   // ---------------------------------
   // Simulation

   // IO-mapping for the valves most be commented-out, to make simulation work.
   #motorValveSimulation_1(speed := #speed, io := #valve1.hmi.io);
   #motorValveSimulation_2(speed := #speed, io := #valve2.hmi.io);
END_FUNCTION_BLOCK

FUNCTION_BLOCK "pulsValve"   // FB13, SCL
{ S7_Optimized_Access := 'TRUE' }
VERSION : 0.1
   VAR_INPUT
      iOpening : Bool;
      iCloses : Bool;
      iPuls : Bool;
      iFullyOpen : Bool;
      iFullyClosed : Bool;
      iConfTimeout : Time := T#3S;
      iConfPulsesBetweenOpenAndClosed : Int;
   END_VAR
   VAR_OUTPUT
      qPos : Real;
      qUnknownPos : Bool;
   END_VAR
   VAR
      cnt : Int;
      rtrig_puls : R_TRIG;
      "timer" : IEC_TIMER;
      first_scan : Bool := TRUE;
   END_VAR
   VAR CONSTANT
      NUMBER_PULES_NOT_CONFIGERED : Int := 0;
   END_VAR
BEGIN
   // Valve position based on puls feedback 

   #rtrig_puls(CLK := #iPuls);
   #"timer".TON(IN := (#iOpening OR #iCloses) AND NOT #rtrig_puls.Q,
              PT := #iConfTimeout);
   IF #iConfPulsesBetweenOpenAndClosed = 0 // Number of pules not configured
       OR #"timer".Q
       OR #first_scan  // 
   THEN
       #qUnknownPos := true;
   ELSIF #iFullyOpen THEN
       #cnt := #iConfPulsesBetweenOpenAndClosed;
       #qUnknownPos := false;
   ELSIF #iFullyClosed THEN
       #cnt := 0;
       #qUnknownPos := false;
   ELSE
       IF #iOpening AND #iCloses THEN
           ; // No action
       ELSIF #rtrig_puls.Q THEN
           #cnt += BOOL_TO_INT(#iOpening);
           #cnt -= BOOL_TO_INT(#iCloses);
       END_IF;
   END_IF;
   #qPos := INT_TO_REAL(#cnt) / INT_TO_REAL(#iConfPulsesBetweenOpenAndClosed) * 100;
   #first_scan := false;
END_FUNCTION_BLOCK

FUNCTION_BLOCK "_loadBalancer_example"   // FB14, SCL
{ S7_Optimized_Access := 'TRUE' }
VERSION : 0.1
   VAR
      load_balancer : "loadBalancer";
   END_VAR
   VAR RETAIN
      devices : Array[1..3] of "load_balancer_device_udt";
      settings : "load_balancer_settings_udt";   // Comman settings
   END_VAR
   VAR
      ___ : Bool;
      pid_output : Real;
      in_1_available : Bool;
      in_1_in_opreation : Bool;
      in_2_available : Bool;
      in_2_in_opreation : Bool;
      in_3_available : Bool;
      in_3_in_opreation : Bool;
      out_1 : Bool;
      out_2 : Bool;
      out_3 : Bool;
      out_1_value : Real;
      out_2_value : Real;
      out_3_value : Real;
   END_VAR
BEGIN
   // Load balancer example:

   // - If devices (eg. pumps) work in parallell, the function will add
   //   or remove devices to operate as the demand increase or decrease.
   // - For vfd, there should be configured a long enough ramp time to
   //   make a smooth transition when a device is added or removed for
   //   operation.
   // - More devices can be controlled, by expand the #devices array.
   // - For this theoretically example static variables bellow "___"
   //   are used, in real application the static variables would be
   //   fysical io.

   // - IMPORTANT: both #devices and #settings need to be set to retain.

   // Available: Eg. in auto, no emergensy stop, no comm.error, ready, etc.
   #devices[1].available := #in_1_available;
   #devices[2].available := #in_2_available;
   #devices[3].available := #in_3_available;

   // input:     Typically the output of a pid-controller, the "damand".
   // devices:   A array, one element for each device.
   // settings:  Can be connected to faceplate in hmi, 
   #load_balancer(input := #pid_output,
                  devices := #devices,
                  settings := #settings );
   // - Important: both #devices and #settings need to be set to retain.
   // - Open the block to see the description inside.

   // Output to devices.
   #out_1 := #devices[1].Q;
   #out_2 := #devices[2].Q;
   #out_3 := #devices[3].Q;

   // If vfd devices is controll by a vfd, then the pid_output shuld be forwared
   // to the vfd's:    
   #out_1_value := SEL(G := #devices[1].Q, IN0 := 0, IN1 := #pid_output);
   #out_2_value := SEL(G := #devices[2].Q, IN0 := 0, IN1 := #pid_output);
   #out_3_value := SEL(G := #devices[3].Q, IN0 := 0, IN1 := #pid_output);
END_FUNCTION_BLOCK

FUNCTION_BLOCK "analogIn_fb"   // FB18, SCL
{ S7_Optimized_Access := 'TRUE' }
VERSION : 0.1
   VAR_INPUT
      in : Int;
   END_VAR
   VAR RETAIN
      aiUdt : "analogInUdt";
   END_VAR
   VAR
      normX : "normXAnalogUdt";
   END_VAR
BEGIN

   "analogIn"(in := #in, aiUdt := #aiUdt, normX := #normX);
END_FUNCTION_BLOCK

FUNCTION_BLOCK "example_stateMachine"   // FB21, SCL
{ S7_Optimized_Access := 'TRUE' }
VERSION : 0.1
   VAR
      state : Int;
      timer1 : "stateMachineTimer";
      timer2 : "stateMachineTimer";
      __condition_1__ : Bool := TRUE;
      __condition_2__ : Bool := TRUE;
      HMI_status : String[100];
   END_VAR
BEGIN
   // State machine with timer example. (https://github.com/rexhip/)

   CASE #state OF
       0:  // Next state after 14 sec. Note that the timer is only one line of code.
           #state += BOOL_TO_INT("sTimer"(pt := T#14s, t := #timer1));

           #HMI_status := CONCAT(IN1 := 'State 0, remaining time: ',
                                 IN2 := "::"(in := #timer1.rt), IN3 := '.');

       1:  // Next state after 7 sec, and '__condition_1__' is true.
           #timer1.pt := T#7s;
           #state += BOOL_TO_INT(#timer1.q AND #__condition_1__);

           // Back to stae 0 if 50 sec elapses. A timer can be used once in each state,
           // therfor timer2 used for this condition. Note the ":=" and not "+=" as above.
           #state := SEL(G := "sTimer"(pt := T#1m50s, t := #timer2), IN0 := #state, IN1 := 0);

           #HMI_status := CONCAT(IN1 := 'State 1, Timer1 ', IN2 := "::"(in := #timer1.rt),
                                 IN3 := ', Timer2 ', IN4 := "::"(in := #timer2.rt));

       2:  // Back to state 0, when '__condition_2__' has been true for 8 sec continuously.
           // The sTimer FC could have been used here also, but for the sake of the
           // example it isn't.
           IF #__condition_2__ THEN
               #timer1.pt := T#8s;
               #state := SEL(G := #timer1.q, IN0 := #state, IN1 := 0);
           END_IF;

           #HMI_status := 'State 2.';
   END_CASE;

   #timer1(state := #state); // Run the timer code.
   #timer2(state := #state);
END_FUNCTION_BLOCK

FUNCTION_BLOCK "modbus_test_rtu_1500"   // FB102, SCL
{ S7_Optimized_Access := 'TRUE' }
VERSION : 0.1
   VAR
      mb_master_1500_ctrl : "mb_master_1500_ctrl";
      mb_query : "mb_query";
      temperature_1 : "Jdrk_RS_WS_N01_8";
      temperature_2 : "Jdrk_RS_WS_N01_8";
      temperature_3 : "Jdrk_RS_WS_N01_8";
      sb_temp_no_answer_1 : "sb_temp_no_answer";
      sb_temp_no_answer_2 : "sb_temp_no_answer";
      sb_temp_no_answer_3 : "sb_temp_no_answer";
      sb_temp_error_1 : "sb_temp_error";
      sb_temp_error_2 : "sb_temp_error";
      sb_temp_error_3 : "sb_temp_error";
      delay_between_queries : "mb_delay_between_queries";
      mb_delay : "mb_delay";
   END_VAR
BEGIN

   #mb_master_1500_ctrl.conf.parity := 0;
   #mb_master_1500_ctrl(hardware_id := 269,
                        operating_mode := 4,
                        baud := 9600,
                        mb_query := #mb_query);

   #delay_between_queries(mb_query := #mb_query);


   #temperature_1(mb_query := #mb_query);
   #temperature_2(mb_query := #mb_query);
   #temperature_3(mb_query := #mb_query);

   #mb_delay(mb_query := #mb_query);

   #sb_temp_no_answer_1(mb_query := #mb_query);
   #sb_temp_no_answer_2(mb_query := #mb_query);
   #sb_temp_no_answer_3(mb_query := #mb_query);

   #sb_temp_error_1(mb_query := #mb_query);
   #sb_temp_error_2(mb_query := #mb_query);
   #sb_temp_error_3(mb_query := #mb_query);
END_FUNCTION_BLOCK

FUNCTION "movingAverageFilter" : Void   // FC1, SCL
{ S7_Optimized_Access := 'TRUE' }
VERSION : 0.1
   VAR_INPUT
      in : Real;
   END_VAR
   VAR_IN_OUT
      filterConst : Real;   // 0=off.
      Q : Real;
   END_VAR
   VAR_TEMP
      z : LReal;
   END_VAR
BEGIN
   // Running average smoothing filter.
   //  - Filter constant has to greater then zero
   //  - PLC scan time will affect the filter.

   IF #filterConst = 0 THEN // Zero -> disable filter 
       #Q := #in;
   ELSE
       #filterConst := MAX(IN1 := 0, IN2 := #filterConst);
       // Creating a number betwwen zero and less then one.
       #z := -1 / REAL_TO_LREAL(#filterConst + 1); 
       #Q := LREAL_TO_REAL(#z * REAL_TO_LREAL(#Q)
                           + (1 - #z) * REAL_TO_LREAL(#in));
   END_IF;
END_FUNCTION

FUNCTION "real2time_format" : Time   // FC1, SCL
{ S7_Optimized_Access := 'TRUE' }
VERSION : 0.1
   VAR_INPUT
      in : Real;
      format : SInt;   // 1=ms, 2=sec, 3=min, 4=h, 5=day
   END_VAR
BEGIN
   // PT-max: 24 days, 20 hours, 31 min, 23 sec and 647 ms.

   // Format: 1=ms, 2=sec, 3=min, 4=h, 5=day

   #real2time_format := T#0s;
   CASE #format OF
       1:  // ms
           #real2time_format := T_CONV(REAL_TO_DINT(#in));
       2:  // Sec
           #real2time_format := T_CONV(REAL_TO_DINT(#in * 1000));
       3:  // Min
           #real2time_format := T_CONV(REAL_TO_DINT(#in * 60000)); //  1000*60
       4:  // Hours
           #real2time_format := T_CONV(REAL_TO_DINT(#in * 3600000)); // 1000*60*60
       5:  // Days
           #real2time_format := T_CONV(REAL_TO_DINT(#in * 86400000)); // 1000*60*60*24
   END_CASE;
END_FUNCTION

FUNCTION "time2real_format" : Real   // FC2, SCL
{ S7_Optimized_Access := 'TRUE' }
VERSION : 0.1
   VAR_INPUT
      in : Time;
      format : SInt;   // 1=ms, 2=sec, 3=min, 4=h, 5=day
   END_VAR
BEGIN
   // PT-max: 24 days, 20 hours, 31 min, 23 sec and 647 ms.

   // Format: 1=ms, 2=sec, 3=min, 4=h, 5=day

   #time2real_format := 0;
   CASE #format OF
       1:  // ms
           #time2real_format := DINT_TO_REAL(T_CONV(#in));
       2:  // Sec
           #time2real_format := DINT_TO_REAL(T_CONV(#in)) / 1000;
       3:  // Min
           #time2real_format := DINT_TO_REAL(T_CONV(#in)) / 60000; // 1000*60
       4:  // Hours
           #time2real_format := DINT_TO_REAL(T_CONV(#in)) / 3600000; // 1000*60*60
       5:  // Days
           #time2real_format := DINT_TO_REAL(T_CONV(#in)) / 86400000; // 1000*60*60*24
   END_CASE;
END_FUNCTION

FUNCTION "analogIn" : Void   // FC4, SCL
TITLE = Analog input
{ S7_Optimized_Access := 'TRUE' }
VERSION : 0.1
   VAR_INPUT
      in : Int;
   END_VAR
   VAR_IN_OUT
      aiUdt : "analogInUdt";
      normX : "normXAnalogUdt";
   END_VAR
   VAR_TEMP
      u : Real;
      x : Real;
      y : Real;
      "e" : Int;
   END_VAR
BEGIN
   // Analog input scaling.

   #u := NORM_X(MIN := #normX.rawMin, VALUE := #in, MAX := #normX.rawMax);
   "movingAverageFilter"(in := #u,
                         filterConst := #aiUdt.filterConst,
                         Q := #aiUdt.unitInterval);
   IF #aiUdt.sim THEN
       ; // A simulated value can be set directly to #aiUdt.Q and #aiUdt.Error
   ELSE
       // Scale back up to raw-value to check if outside error limits.
       #x := SCALE_X(MIN := #normX.rawMin, MAX := #normX.rawMax,
                     VALUE := #aiUdt.unitInterval);
       #aiUdt.Error := #x < #normX.errorLimMin OR #x > #normX.errorLimMax;
       // Log the time when the error occurred.
       IF #aiUdt.Error AND NOT #aiUdt.zOldError THEN
           #"e" := RD_LOC_T(#aiUdt.ErrorTime);
       END_IF;

       IF #aiUdt.Error THEN
           #y := SINT_TO_REAL(#aiUdt.errorAction) / 100;
       ELSIF #aiUdt.forceInsideScale THEN
           #y := LIMIT(MN := 0, IN := #aiUdt.unitInterval, MX := 1);
       ELSE
           #y := #aiUdt.unitInterval;
       END_IF;
       #aiUdt.Q := SCALE_X(MIN := #aiUdt.scaleMin, MAX := #aiUdt.scaleMax,
                           VALUE := #y ) * #aiUdt.gain + #aiUdt.offset;
   END_IF;
   #aiUdt.zOldError := #aiUdt.Error;

   // ( https://github.com/rexhip/ )
END_FUNCTION

FUNCTION "boost_start" : Void   // FC5, SCL
{ S7_Optimized_Access := 'TRUE' }
VERSION : 0.1
   VAR_INPUT
      t_diff : USInt;
      start : Bool;
   END_VAR
   VAR_OUTPUT
      reset_timers : Bool;
   END_VAR
   VAR_IN_OUT
      devices : Array[*] of "load_balancer_device_udt";
      settings : "load_balancer_settings_udt";
      info : "load_balancer_info_udt";
      boost_start : SInt;
      set : SInt;
   END_VAR
   VAR_TEMP
      c : DInt;
      u : DInt;
      lower : DInt;
   END_VAR
BEGIN
   #lower := LOWER_BOUND(ARR := #devices, DIM := 1);
   FOR #c := #lower TO UPPER_BOUND(ARR := #devices, DIM := 1) DO

       #u := #c - #lower + 1; // #u start at 1, increasing by 1 for each iteration.
       IF #settings.boostStart.reset THEN
           // Reset stastic, on how many devices is operating same time.
           #devices[#c].z.n_cnt := 0;
       ELSIF #settings.info.started = #u THEN
           // Log how many devices is operating same time, most fequently.
           #devices[#c].z.n_cnt += #t_diff;
       END_IF;

       // Change how many devices to boost start at startup, based on how many
       // devices is most commenly used.
       IF #settings.boostStart.auto
           AND #devices[#c].z.n_cnt >
           (* *)#devices[#lower + #settings.boostStart.devices - 1].z.n_cnt
       THEN
           #settings.boostStart.devices := DINT_TO_USINT(#u);
       END_IF;
   END_FOR;

   // Set a number of operating devices. (Without waiting for the input and the timers)
   IF #set > -1 THEN
       #boost_start := #set - UINT_TO_SINT(#info.devices_started);

       // Do boost start when input change away from zero.    
   ELSIF #settings.boostStart.enable // HMI enable.
       AND #start
       AND #set = -1
   THEN
       #boost_start :=
       UINT_TO_SINT(#settings.boostStart.devices - #info.devices_started);
   END_IF;
   // #set is put back to -1 at the bottom of the block.

   // MN: Devies started to be stopped.
   // MX: Devices available for start. 
   #boost_start := LIMIT(MN := - UINT_TO_SINT(#info.devices_started),
                         IN := #boost_start,
                         MX := UINT_TO_SINT(#info.devices_standby));

   #reset_timers := #boost_start <> 0 OR #set <> -1; // Reset timers.
END_FUNCTION

FUNCTION "analogInReal" : Void   // FC7, SCL
{ S7_Optimized_Access := 'TRUE' }
VERSION : 0.1
   VAR_INPUT
      in : Real;
      error : Bool;
   END_VAR
   VAR_IN_OUT
      aiUdt : "analogInAndAlarmsUdt";
      ioGlobal : "ioGlobal_FB";
   END_VAR
   VAR_TEMP
      dommy : Int;
      u : Real;
   END_VAR
BEGIN
   // Analog input 
   // Wrapper to use analog input block with real input.
   // 
   #aiUdt.ai.Error := #error;

   IF #aiUdt.ai.sim THEN
       ; // A simultated value may be set directly at: #ai.ai.Q
   ELSE
       #u := #in * #aiUdt.ai.gain + #aiUdt.ai.offset;
       "movingAverageFilter"(in := #u,
                             filterConst := #aiUdt.ai.filterConst,
                             Q := #aiUdt.ai.Q);
   END_IF;

   #aiUdt.execAiLogic := false;
   "analogInAndAlarms"(in := #dommy,
                       aiUdt := #aiUdt,
                       ioGlobal := #ioGlobal);

   // ( https://github.com/rexhip/ )
END_FUNCTION

FUNCTION "analogOut" : Void   // FC9, SCL
{ S7_Optimized_Access := 'TRUE' }
VERSION : 0.1
   VAR_OUTPUT
      q : Int;
   END_VAR
   VAR_IN_OUT
      aoUdt : "analogOutUdt";
      ioGlobal : "ioGlobal_FB";
   END_VAR
   VAR_TEMP
      x : Real;
      y : Real;
   END_VAR
BEGIN
   // Analog out 

   // - failSafe: Output will go to a predefined value set by
   //   failSafeValue (%), this can be used for emergency stop.
   //   Simulation will not work when failSafe is activated.

   // A id for each io
   #ioGlobal.z.ioIdCnt += 1;

   IF #ioGlobal.info2ioBlocks.disableAllSim THEN
       #aoUdt.simEnable := false;
   END_IF;

   IF #aoUdt.failSafe THEN
       #x := SINT_TO_REAL(#aoUdt.failSafeValue) / 100 ; // [%]
   ELSE
       IF #aoUdt.simEnable THEN
           #y := #aoUdt.simValue;
       ELSIF #aoUdt.interlook THEN
           #y := 0;
       ELSE
           #y := #aoUdt.in;
       END_IF;
       #x := NORM_X(MIN := #aoUdt.scaleMin, VALUE := #y,
                    MAX := #aoUdt.scaleMax);
       #aoUdt.simValue := #y;
   END_IF;
   #x := LIMIT(MN := 0, IN := #x, MX := 1);
   #q := SCALE_X(MIN := #ioGlobal.normX.rawMin, VALUE := #x,
                     MAX := #ioGlobal.normX.rawMax);

   #ioGlobal.collectInfo.activeSimCnt += BOOL_TO_UINT(#aoUdt.simEnable);

   // ( https://github.com/rexhip/ )
END_FUNCTION

FUNCTION "ioGlobalMotorValveLinking" : Void   // FC24, SCL
{ S7_Optimized_Access := 'TRUE' }
VERSION : 0.1
   VAR_IN_OUT
      ioGlobal : "ioGlobal_FB";
      valve : "motorValve";
   END_VAR
BEGIN
   // Link ioGlobal with valve functions.

   // A id for each io
   #ioGlobal.z.ioIdCnt += 1;

   IF #ioGlobal.info2ioBlocks.disableAllSim THEN
       #valve.hmi.sim.enable := false;
   END_IF;
   // Count active simulations
   #ioGlobal.collectInfo.activeSimCnt +=
   BOOL_TO_UINT(#valve.hmi.sim.enable OR #valve.hmi.sim.simByPlc);

   // Count number of errors
   #ioGlobal.collectInfo.errorCnt +=
   BOOL_TO_UINT(#valve.hmi.io.in.posError OR #valve.hmi.error.timeout);
END_FUNCTION

FUNCTION "real_to_time" : Time   // FC29, SCL
{ S7_Optimized_Access := 'TRUE' }
VERSION : 0.1
   VAR_INPUT
      in : Real;
   END_VAR
BEGIN

   #real_to_time := T_CONV(REAL_TO_DINT(#in * 1000));
END_FUNCTION

// folder: Library/Alternating/Load balancer/Blocks and UDT's

FUNCTION_BLOCK "loadBalancer"   // FB13, SCL
{ S7_Optimized_Access := 'TRUE' }
VERSION : 0.1
   VAR_INPUT
      input : Real;   // [%] Typically a output from a pid-controller.
   END_VAR
   VAR_IN_OUT
      devices : Array[*] of "load_balancer_device_udt";   // Variables for each device.
      settings : "load_balancer_settings_udt";   // Comman settings
   END_VAR
   VAR RETAIN
      conf : Struct   // Advanced configuration
         enable_operation_time_cnt : Bool := true;   // Enable operation time cnt
         at_least_one : Bool := true;   // At least one device will always be in operation
         bypass_InOperation_signal : Bool := true;   // Output control in-operation variable.
         input_zero_reset : Time := T#10M;   // All outputs will be turn off if input has been zero for this time.
         exec_boost_start_code : Bool := true;
      END_STRUCT;
   END_VAR
   VAR
      boost_start : SInt;   // Start a relative number of devices. (Negative number will stop devices)
      set : SInt := -1;   // Start a exact number of devices. (Set back to -1 right away)
      _ : Bool;
      timer_start : IEC_TIMER;
      timer_start_q : Bool;
      timer_stop : IEC_TIMER;
      timer_stop_q : Bool;
      timer_input_zero : IEC_TIMER;
      old_sec : USInt;
      ftrig_zero_input_timer : F_TRIG;
      runtime_mem1 : LReal;
      runtime_mem2 : LReal;
   END_VAR
   VAR_TEMP
      candidates : Struct
         start : Struct
            index : DInt;
            operation_time : UDInt;
         END_STRUCT;
         stop : Struct
            index : DInt;
            operation_time : UDInt;
         END_STRUCT;
      END_STRUCT;
      info : "load_balancer_info_udt";
      lower : DInt;
      upper : DInt;
      c : DInt;
      t_diff : USInt;
      oper : SInt;
      u : DInt;
      reset_timers : Bool;
      dommy : Bool;
   END_VAR
   VAR CONSTANT
      NO_CANDIDATE : DInt := 16#7fffffff;
   END_VAR
BEGIN
   (* === Load balancer ===    

   - If devices (eg. pumps) work in parallell, the function will start or stop devices
     to operate as the demand increase or decrease.
   - A devices will be added for operation, if #input is above a certain value for a
     ceratin time, eg above 90% for 50 seconds. Likewise a devices will be removed from
     operation if #input is bellow a certain value for a certain time, eg. 10% for 30
     secunds. The limits and the times are adjustable inside #settings.
   - It's the device with least operating time that will be added first, and the device
     with most operating hours will be removed from operation first.
   - #input will typically be the output of a pid-controller.
   - For vfd, there should be configured a ramp time to make a smooth transition when a
     device is added or removed for operation.
   - #devices[*].in.in_operation, is a input for fyscical feedback signal from the
     devices. this feature can be disabled by setting
     #load_balancer.conf.bypass_InOperation_signal, to true.
   - #boost_start: Make more then one devices start right away, without have to wait for
     them to start one by one. Use a negative number to stop several devies at once. One
     scan is need to start or stop each device.
   - #set: Will start or stop devies to mache number of the variable. This block will set
     the variable to -1 for the next scan.

   *)

   // If input is zero for a certain time, then all outputs is set to false.
   #timer_input_zero.TON(IN := #input = 0, PT := #conf.input_zero_reset);
   // Used to set correct number of devices from start. (Boost start)
   #ftrig_zero_input_timer(CLK := NOT #timer_input_zero.Q);

   // Default values, if the value isn't overwritten after the
   // for-loop (bellow), then there is "no candidate".
   #candidates.stop.index := #NO_CANDIDATE;
   #candidates.start.index := #NO_CANDIDATE;
   // Set to max, try find a lesser value in the for-loop bellow.
   #candidates.start.operation_time := 16#ffffffff;

   // Operating time preparing calculations:
   #runtime_mem2 += RUNTIME(#runtime_mem1);
   #t_diff := LREAL_TO_USINT(FLOOR(#runtime_mem2)); // "Overflow" if >= 1 sec.
   #runtime_mem2 -= USINT_TO_LREAL(#t_diff);

   // Boost start makes, more then one device start right away.
   IF #conf.exec_boost_start_code THEN
       "boost_start"(t_diff := #t_diff,
                     start := #ftrig_zero_input_timer.Q,
                     reset_timers => #reset_timers,
                     devices := #devices,
                     settings := #settings,
                     info := #info,
                     boost_start := #boost_start,
                     set := #set);
   END_IF;

   #lower := LOWER_BOUND(ARR := #devices, DIM := 1);
   #upper := UPPER_BOUND(ARR := #devices, DIM := 1);
   FOR #c := #lower TO #upper DO

       #devices[#c].Q := #devices[#c].Q
       (* *)AND #devices[#c].available // Disable devices that are not available. 
       (* *)AND NOT #timer_input_zero.Q // Input has not been zero for a ceratain time.
       OR #settings.bypass; // If bypass, then enable all devices.

       // If no fysical feedback signal from device for "in-operation", then
       // it's possible to bypass it.
       IF #conf.bypass_InOperation_signal THEN
           #devices[#c].in_operation := #devices[#c].Q;
       END_IF;

       REGION Candidates        
           // Candidate device to be stoped (the one that has the longest operating time)
           IF #devices[#c].Q // In use
               AND #devices[#c].operation_time >= #candidates.stop.operation_time
           THEN
               #candidates.stop.index := #c;
               #candidates.stop.operation_time := #devices[#c].operation_time;
           END_IF;

           // Candidate device to be started (the one that has the least operating time)
           IF #devices[#c].available
               AND NOT #devices[#c].Q // not allready in use
               AND #devices[#c].operation_time < #candidates.start.operation_time
           THEN
               #candidates.start.index := #c;
               #candidates.start.operation_time := #devices[#c].operation_time;
           END_IF;
       END_REGION

       REGION Collect-statistics
           // Operating time cnt. (#t_diff will always be zero, if the feature is disabled)
           #devices[#c].operation_time += SEL(G := #devices[#c].in_operation
                                              AND #conf.enable_operation_time_cnt,
                                              IN0 := 0, IN1 := USINT_TO_UDINT(#t_diff));
           // Count number of devices in operation.
           #info.devices_in_operation += BOOL_TO_UINT(#devices[#c].in_operation);
           // Count number of devices in standby.
           #info.devices_standby +=
           BOOL_TO_UINT(#devices[#c].available
                        AND NOT #devices[#c].Q); // NOT #devices[#c].in.in_operation
           // Count number of devices started.
           #info.devices_started += BOOL_TO_UINT(#devices[#c].Q);
       END_REGION
   END_FOR;

   // Some info (for hmi)
   #settings.info.total := DINT_TO_UINT(#upper - #lower + 1);

   // If for some reason, the number operating devies can be limited to less
   // then available
   #settings.max_devices_same_time := // A setting.
   LIMIT(MN := 1,
         IN := #settings.max_devices_same_time,
         MX := #settings.info.total);

   // Force min value for param.
   #settings.max_diff_operating.sec :=
   MAX(IN1 := 60, IN2 := #settings.max_diff_operating.sec);

   // Timers for adding and removing devices for operation.

   #timer_stop.TON(IN := #input < #settings.stop.limit AND NOT #reset_timers,
                   PT := #settings.stop.delay,
                   Q => #timer_stop_q);
   #timer_start.TON(IN := #input > #settings.start.limit AND NOT #reset_timers,
                    PT := #settings.start.delay,
                    Q => #timer_start_q);

   REGION start-stopp
       // Stoping a device
       IF NOT #settings.bypass // The bypass-function turn on all outputs. 
           AND #candidates.stop.index <> #NO_CANDIDATE // A device is available 
           AND (#info.devices_in_operation > 1 // Can't remove last device in operation
           (* *)OR NOT #conf.at_least_one)  // Possible to disable the feature
           AND (
           (* *)#info.devices_in_operation > #settings.max_devices_same_time
           (* *)OR #timer_stop_q // If #input below a certain value for a certain time
           (* *)OR #settings.stop.force  // Used to stop the next device (hmi)
           (* *)OR #boost_start < 0)
       THEN
           #devices[#candidates.stop.index].Q := false; // Disable one device
           RESET_TIMER(#timer_stop);
           #oper := -1;
           // Increase var until zero.
           #boost_start := SEL(G := #boost_start < 0, IN0 := 0, IN1 := #boost_start + 1);

           // Start a devices.
       ELSIF #candidates.start.index <> #NO_CANDIDATE // A device is available 
           AND #info.devices_in_operation < #settings.max_devices_same_time
           AND #input > 0 AND (
           (* *)#info.devices_in_operation < 1 // At least one device operating
           (*      *)AND #conf.at_least_one // Possible to disable the feature
           (* *)OR #timer_start_q // If #input above a certain value for a certain time
           (* *)OR #settings.start.force // Used to starp the next device (hmi)
           (* *)OR #boost_start > 0)
       THEN
           #devices[#candidates.start.index].Q := true; // Enable one more device
           RESET_TIMER(#timer_start);
           #oper := 1;
           // Decrease var until zero.
           #boost_start := SEL(G := #boost_start > 0, IN0 := 0, IN1 := #boost_start - 1);

           // Change operating device, if the operating-time between two devies is to large.
       ELSIF #settings.max_diff_operating.enable
           AND #candidates.start.index <> #NO_CANDIDATE // A candidate is available to be started
           AND #candidates.stop.index <> #NO_CANDIDATE // A candidate is available to be stoped
           AND (#candidates.stop.operation_time - #candidates.start.operation_time >
           (* *)#settings.max_diff_operating.sec) // And the difference is to large.
       THEN
           // Stop the device with most operating time and start the devices with
           // least operating time.
           #devices[#candidates.stop.index].Q := false;
           #devices[#candidates.start.index].Q := true;
       END_IF;
   END_REGION

   // Update vars, after start or stop a device. (above)
   #info.devices_in_operation += SINT_TO_UINT(#oper);
   #info.devices_started += SINT_TO_UINT(#oper);
   #info.devices_standby -= SINT_TO_UINT(#oper);

   // Transfer values to hmi-vars
   #settings.info.in_operation := #info.devices_in_operation;
   #settings.info.started := #info.devices_started;
   #settings.info.standby := #info.devices_standby;

   #settings.info.input := #input;

   // Information has been recived, so now back to default values.
   #set := -1;
   #settings.start.force := false;
   #settings.stop.force := false;
   #settings.boostStart.reset := false;

   // https://github.com/rexhip/
END_FUNCTION_BLOCK

// folder: Library/IO-handeling/Analog in/Blocks

FUNCTION "analogInAndAlarms" : Void   // FC6, SCL
{ S7_Optimized_Access := 'TRUE' }
VERSION : 0.1
   VAR_INPUT
      in : Int;
   END_VAR
   VAR_IN_OUT
      aiUdt : "analogInAndAlarmsUdt";
      ioGlobal : "ioGlobal_FB";
   END_VAR
   VAR CONSTANT
      VALUE_LESS_THEN_LIM : SInt := 1;
      VALUE_GREATER_THEN_LIM : SInt := 2;
   END_VAR
BEGIN
   // Analog input with alarm handling. 

   REGION Input handling
       // A id for each io
       #ioGlobal.z.ioIdCnt += 1;

       // Disable all simulations.
       #aiUdt.ai.sim := #aiUdt.ai.sim AND NOT #ioGlobal.info2ioBlocks.disableAllSim;

       IF #aiUdt.execAiLogic THEN // Execute analog input logic
           "analogIn"(in := #in,
                      aiUdt := #aiUdt.ai,
                      normX := #ioGlobal.normX);
       END_IF;
       // Count number of errors
       #ioGlobal.collectInfo.errorCnt += BOOL_TO_UINT(#aiUdt.ai.Error);;
       // Count active simulations 
       #ioGlobal.collectInfo.activeSimCnt += BOOL_TO_UINT(#aiUdt.ai.sim);
   END_REGION

   REGION Alarms  
   // Connecting ioGlobal functions with each alarm.
   "ioGlobalAlarmLinking"(alarm := #aiUdt.alarmHH, ioGlobal := #ioGlobal);
   "ioGlobalAlarmLinking"(alarm := #aiUdt.alarmH, ioGlobal := #ioGlobal);
   "ioGlobalAlarmLinking"(alarm := #aiUdt.alarmLL, ioGlobal := #ioGlobal);
   "ioGlobalAlarmLinking"(alarm := #aiUdt.alarmL, ioGlobal := #ioGlobal);

   "alarmReal"(value := #aiUdt.ai.Q, // HH alarm
               action := #VALUE_GREATER_THEN_LIM,
               disable := false,
               runtimeDiff := #ioGlobal.info2ioBlocks.runtimeDiff,
               alarm := #aiUdt.alarmHH);
   "alarmReal"(value := #aiUdt.ai.Q,// H alarm
               action := #VALUE_GREATER_THEN_LIM,
               disable := #aiUdt.alarmHH.Q,
               runtimeDiff := #ioGlobal.info2ioBlocks.runtimeDiff,
               alarm := #aiUdt.alarmH);
   "alarmReal"(value := #aiUdt.ai.Q, // LL alarm
               action := #VALUE_LESS_THEN_LIM,
               disable := false,
               runtimeDiff := #ioGlobal.info2ioBlocks.runtimeDiff,
               alarm := #aiUdt.alarmLL);
   "alarmReal"(value := #aiUdt.ai.Q, // L alarm
               action := #VALUE_LESS_THEN_LIM,
               disable := #aiUdt.alarmLL.Q,
               runtimeDiff := #ioGlobal.info2ioBlocks.runtimeDiff,
               alarm := #aiUdt.alarmL);
   END_REGION

   REGION HMI-features
       // Copy paste all settings. (HMI)
       IF #aiUdt.hmi.copyAllSettings THEN
           #ioGlobal.copyPaste := #aiUdt;
           #aiUdt.hmi.copyAllSettings := false;
       ELSIF #aiUdt.hmi.pasteAllSettings THEN
           "pasteAnalogInSetting"(src := #ioGlobal.copyPaste, dest := #aiUdt);
           #aiUdt.hmi.pasteAllSettings := false;
       END_IF;

       #aiUdt.hmi.showTag := #ioGlobal.hmi.hmiShowTags;
   END_REGION

   // ( https://github.com/rexhip/ )
END_FUNCTION

FUNCTION "analogInSimple" : Real   // FC13, SCL
{ S7_Optimized_Access := 'TRUE' }
VERSION : 0.1
   VAR_INPUT
      mn : Real;
      in : Int;
      mx : Real;
   END_VAR
   VAR_TEMP
      x : Real;
   END_VAR
BEGIN
   // Analog in 

   #x := NORM_X(MIN := 0, VALUE := #in, MAX := 27648);
   #x := LIMIT(MN := 0, IN := #x, MX := 1);
   #analogInSimple := SCALE_X(MIN := #mn, VALUE := #x, MAX := #mx);

   // ( https://github.com/rexhip/ )
END_FUNCTION

// folder: Library/Modbus/.Start examples

FUNCTION_BLOCK "modbus_rtu_1500"   // FB5, SCL
{ S7_Optimized_Access := 'TRUE' }
VERSION : 0.1
   VAR
      mb_query : "mb_query";
      mb_master_1500_ctrl : "mb_master_1500_ctrl";
      abb_aquaMaster_device1 : "abb_aquaMaster_3";
      abb_aquaMaster_device2 : "abb_aquaMaster_3";
      abb_aquaMaster_device3 : "abb_aquaMaster_3";
      resault_data_1 : Word;
   END_VAR
BEGIN
   // hardware_id:     May be found inside the hardware configuration.
   // operating_mode:  0: RS232, 2: RS422, 4: RS485.
   // baud:            Bits per sec. (Parity is even by default)
   // timeout:         Automatically calculated if set to zero. (T#0s)
   // mb_query:        The FB that connects everything together.
   #mb_master_1500_ctrl(hardware_id := 0, // REPLACE WITH CORRECT ID.
                        operating_mode := 4, // RS-485
                        baud := 19200, // bps
                        mb_query := #mb_query);

   // Each blocks bellow represent one device on the bus. 
   #abb_aquaMaster_device1(mb_addr := 1, mb_query := #mb_query);
   #abb_aquaMaster_device2(mb_addr := 2, mb_query := #mb_query);
   #abb_aquaMaster_device3(mb_addr := 3, mb_query := #mb_query);


   // Debugging tip, (no code)
   "mb_Debugging"();
END_FUNCTION_BLOCK

FUNCTION_BLOCK "modbus_tcp"   // FB79, SCL
{ S7_Optimized_Access := 'TRUE' }
VERSION : 0.1
   VAR
      mb_query : "mb_query";
      mb_client_ctrl : "mb_client_ctrl";
      siemens_PAC3200 : "siemens_PAC3200";
      ip : Array[1..4] of Byte;
      mb_delay_between_queries : "mb_delay_between_queries";
   END_VAR
BEGIN
   // IP-address of the modbus server
   #ip[1] := 192;
   #ip[2] := 168;
   #ip[3] := 1;
   #ip[4] := 2;

   // interface:  Profinet interface.
   //             (Find const. inside "Device configuration")
   // conn_id:    A unique id for each tcp connectin in the plc.
   // ip_addr:    The ip-address of the server. (Array of 4 bytes)
   // tcp_port:   Default port is 502. (UDP isn't available)
   // timeout:    Depends on the network conncetion.
   // mb_query:   The query FB.
   #mb_client_ctrl(interface := 0, // REPLACE WITH CORRECT ID OR CONST,
                                   // Eg. "Local~PROFINET_interface_1",
                   conn_id := 123,
                   ip_addr := #ip,
                   tcp_port := 502,
                   timeout := T#400ms,
                   mb_query := #mb_query);

   // Delay the query execution, this prevent the plc from
   // jamming the network. Adjust the time to the application.
   #mb_delay_between_queries(delay := T#500ms,
                             mb_query := #mb_query);

   #siemens_PAC3200(mb_query := #mb_query);


   // Debugging tip, (no code)
   "mb_Debugging"();
END_FUNCTION_BLOCK

FUNCTION_BLOCK "modbus_rtu_1200"   // FB98, SCL
{ S7_Optimized_Access := 'TRUE' }
VERSION : 0.1
   VAR
      mb_query : "mb_query";
      mb_master_1200_ctrl : "mb_master_1200_ctrl";
      abb_aquaMaster_device1 : "abb_aquaMaster_3";
      abb_aquaMaster_device2 : "abb_aquaMaster_3";
      abb_aquaMaster_device3 : "abb_aquaMaster_3";
      Auma_valve : "Auma_valve";
      Phoenix_Contact_UPS : "Phoenix_Contact_UPS";
      resault_data_1 : Word;
      Phoenix_Contact_UPS_1 : "Phoenix_Contact_UPS";
   END_VAR
BEGIN
   // hardware_id: Can be found inside "Device configuration".
   // baud:        Bits per sec. (Parity is even by default)
   // timeout:     Automatically calculated if set to T#0s.
   // mb_query:    The FB that connects everything together.
   #mb_master_1200_ctrl(hardware_id := 0, // REPLACE WITH CORRECT ID.
                        baud := 19200,
                        mb_query := #mb_query);

   // Each blocks bellow represent one device on the bus.

   // Three Abb aqua-master's.
   #abb_aquaMaster_device1(mb_addr := 1, mb_query := #mb_query);
   #abb_aquaMaster_device2(mb_addr := 2, mb_query := #mb_query);
   #abb_aquaMaster_device3(mb_addr := 3, mb_query := #mb_query);

   // A valve 
   #Auma_valve(mb_addr := 4, mb_query := #mb_query);

   // A UPS.
   #Phoenix_Contact_UPS(mb_addr := 5, mb_query := #mb_query);

   // A station block can be used both for both modbus rtu and tcp. This
   // is particular useful if a tcp-rtu-gateway is used. The same program
   // could be used, just swap mb_master_1200_ctrl, with mb_client_ctrl.

   // Read holding register 456 from device with modbus address 123.
   // This is an example showing that a query does not necessarily need
   // to be part of a station block (SB) as obove, however making
   // reusable SB's is good practice.
   #mb_query(mb_addr := 123,
             mode := #mb_query.c.read.holding_reg,
             data_addr := 456,
             data_ptr := #resault_data_1);


   // Debugging tip, (no code)
   "mb_Debugging"();
END_FUNCTION_BLOCK

FUNCTION "mb_Readme" : Void   // FC13, SCL
{ S7_Optimized_Access := 'TRUE' }
VERSION : 0.1
BEGIN
   (* Instructions:

   - Add one of the exmple FB's to your PLC.
   - Call that FB from a cyclic OB.
   - Terminate connection to type on the example FB. (Right click the FB)
   - Set hardware_id, buad-rate, ip, tcp-port, etc, to the correct value.
   - Look inside the library and check if there is a ready station block (SB),
     for your program. If there isn't then a new has to be made. 
   - Station blocks can be single-DB's or multi-instances in a FB.
   - Remove the exmple code and example SB's.

   IMPORTANT: As stated above, the start examples fb, need to be terminated 
              from it's type. If the type is edited and later there is a 
              library update, then all the changes will get lost.

   - Instructions need to be of the latest version, 
     this is usually already set:
     * Instructions -> Communication -> Others -> Modbus TCP
     * Instructions -> Communication -> Communication processor -> Modbus
     * Instructions -> Communication -> Communication processor -> Modbus (RTU)  
     * Instructions -> Basic instructions -> Word logic operations -> SEL.
     Change version in the right column.

   *)
END_FUNCTION

// folder: Library/Modbus/.Start examples/Other start examples

FUNCTION_BLOCK "LAD_modbus_rtu"   // FB97, LAD
TITLE = Example modbus rtu
{ S7_Optimized_Access := 'TRUE' }
VERSION : 0.1
// REPLACE hardware_id WITH CORRECT ID.
   VAR
      mb_master_ctrl : "mb_master_1200_ctrl";
      mb_query : "mb_query";
      aquaMaster_device1 : "abb_aquaMaster_3";
      aquaMaster_device2 : "abb_aquaMaster_3";
      Auma_valve : "Auma_valve";
      Phoenix_Contact_UPS : "Phoenix_Contact_UPS";
   END_VAR
   VAR_TEMP   // added for the SCL form of the ladder/FBD networks
      _w1 : Bool;
   END_VAR
BEGIN

REGION Network 1: Modbus master
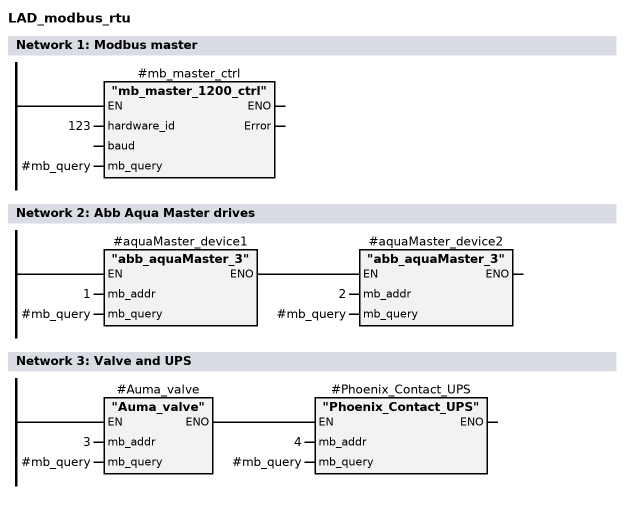
   RUNG wire#powerrail
      #mb_master_ctrl(hardware_id := 123, baud :=, mb_query := #mb_query, Error =>)
   END_RUNG
   // the same network as SCL:
   #mb_master_ctrl(hardware_id := 123, mb_query := #mb_query);   // "mb_master_1200_ctrl"
END_REGION

REGION Network 2: Abb Aqua Master drives
   RUNG wire#powerrail
      #aquaMaster_device1(mb_addr := 1, mb_query := #mb_query)
      #aquaMaster_device2(mb_addr := 2, mb_query := #mb_query)
   END_RUNG
   // the same network as SCL:
   #aquaMaster_device1(mb_addr := 1, mb_query := #mb_query, ENO => #_w1);   // "abb_aquaMaster_3"
   IF #_w1 THEN
       #aquaMaster_device2(mb_addr := 2, mb_query := #mb_query);   // "abb_aquaMaster_3"
   END_IF;
END_REGION

REGION Network 3: Valve and UPS
   RUNG wire#powerrail
      #Auma_valve(mb_addr := 3, mb_query := #mb_query)
      #Phoenix_Contact_UPS(mb_addr := 4, mb_query := #mb_query)
   END_RUNG
   // the same network as SCL:
   #Auma_valve(mb_addr := 3, mb_query := #mb_query, ENO => #_w1);   // "Auma_valve"
   IF #_w1 THEN
       #Phoenix_Contact_UPS(mb_addr := 4, mb_query := #mb_query);   // "Phoenix_Contact_UPS"
   END_IF;
END_REGION
END_FUNCTION_BLOCK

// folder: Library/Modbus/Core/Ctrl

FUNCTION_BLOCK "mb_client_ctrl"   // FB9, SCL
{ S7_Optimized_Access := 'TRUE' }
VERSION : 1.0
   VAR_INPUT
      interface : Hw_Any := 64;   // Profinet interface id
      conn_id : Conn_Ouc := 123;   // Connection id. Should be unique between all tcp connections.
      ip_addr : Array[1..4] of Byte;   // IPv4 address.
      tcp_port : UInt := 502;   // TCP port
      timeout : Time := T#2s;
   END_VAR
   VAR_OUTPUT
      Error : Bool;   // error flag with tof timer
   END_VAR
   VAR_IN_OUT
      mb_query : "mb_query";   // udt mb
   END_VAR
   VAR
      conf : Struct   // Configuration that normal shouldn't need to be changed.
         disconnect : Bool := FALSE;
         retries : USInt := 1;
         timeout_connect : Time;   // May be set longer, then the main timeout. T#0s => Use normal timeout.
         disconnect_on_80A3 : Bool := true;
      END_STRUCT;
      client : MB_CLIENT;
      tdiscon : TDISCON;
      tcon_ip_v4 : TCON_IP_v4;
      ton_connect : TON_TIME;
      end : "mb_internal_e";
      connected_least_once : Bool;   // One connection has taken place.
   END_VAR
   VAR_TEMP
      comm_err : Bool;
   END_VAR
   VAR CONSTANT
      INIT_QUERY : USInt := 2;
      EXEC_QUERY : USInt := 3;
      RECIVE_RESUALT : USInt := 4;
   END_VAR
BEGIN
   // Rexhip - Extended modbus library.
   // Please see top section of mb_query for more info.
   //
   // Modbus tcp for S7-1200 and S7-1500.

   REGION Init
       #tcon_ip_v4.InterfaceId := #interface;
       #tcon_ip_v4.ID := #conn_id;
       #tcon_ip_v4.ConnectionType := 11; // tcp
       #tcon_ip_v4.ActiveEstablished := true;
       #tcon_ip_v4.RemoteAddress.ADDR := #ip_addr;
       #tcon_ip_v4.RemotePort := #tcp_port;

       PRESET_TIMER(PT :=
                    SEL(G := #conf.timeout_connect = T#0s
                        OR NOT #connected_least_once,
                        IN0 := #conf.timeout_connect,
                        IN1 := #timeout),
                    TIMER := #ton_connect);
       #ton_connect(IN := NOT #conf.disconnect AND NOT #client.Connected,
                    PT := #ton_connect.PT);
       // - Use #timeout if: #timeout_connect is set to zero, or there has
       //   been a least one connection to the server.
       // - Establing a TCP connection may take long. 
       // - If mb_client does not establish a connection it will not  throw
       //   timeout error. Timeout is handled manually for that case. 

       // Conversion of function codes. 
       IF #mb_query.z.run.state = #INIT_QUERY THEN
           CASE #mb_query.z.q.mode OF
               1..16: // 1..6, 15, 16:
                   #client.MB_MODE := #mb_query.z.q.mode + 100;
                   // Eg. Siemens use 103 for fc 3. (read halding reg)
               200..202:
                   #client.MB_MODE := #mb_query.z.q.mode - 200;
               ELSE
                   #client.MB_MODE := #mb_query.z.q.mode;
           END_CASE;
           #client.MB_Unit_ID := UINT_TO_BYTE(#mb_query.z.q.mb_addr);
           #client.Retries := #conf.retries;
           #mb_query.z.run.state := #EXEC_QUERY; // Next state.
       END_IF;
   END_REGION

   REGION Exec
       // STATUS 16#80A3 : 
       // If a new download has taken place, and this block is re-initialize,
       // then the mb_client block will output the error code saying that:
       // "Attempt being made to re-establish an existing connection." The
       // solution to this problem is to disconnect and then reconnect. It
       // dosen't work to use disconnect input on the mb_client block.
       #tdiscon(REQ := #client.STATUS = 16#80A3 AND #conf.disconnect_on_80A3,
                ID := #conn_id);

       #client.Rcv_Timeout :=
       (* *)UDINT_TO_REAL(T_CONV(#timeout)) * 0.001; // ms to s.
       #client(DISCONNECT := #conf.disconnect OR #tdiscon.BUSY,
               REQ := #mb_query.z.run.state = #EXEC_QUERY
               AND NOT #client.BUSY
               AND NOT #client.DISCONNECT,
               MB_MODE := #client.MB_MODE,
               MB_DATA_ADDR := #mb_query.z.q.data_addr,
               MB_DATA_LEN := #mb_query.z.q.data_len,
               BUSY => #mb_query.stat.busy,
               MB_DATA_PTR := #mb_query.z.buffer,
               CONNECT := #tcon_ip_v4);

       IF #mb_query.z.run.state = #EXEC_QUERY THEN
           #mb_query.stat.error := #client.ERROR OR #ton_connect.Q;
           #mb_query.stat.done := #client.DONE AND NOT #mb_query.stat.error;
           #mb_query.stat.status := #client.STATUS;
           // Comm. error and timeout handeling. 
           CASE WORD_TO_UINT(#mb_query.stat.status) OF
               16#80C8,  // No response from the server.
               16#818C: // blocked_proc_timeout or rcv_timeout.
                   #comm_err := #mb_query.stat.error;
           END_CASE;
           #mb_query.stat.error_comm := #ton_connect.Q OR #comm_err;
       END_IF;
   END_REGION

   // End is a comman FB for both tcp and rtu.
   #end(mb_query := #mb_query, Error => #Error);
END_FUNCTION_BLOCK

FUNCTION_BLOCK "mb_master_1500_ctrl"   // FB10, SCL
{ S7_Optimized_Access := 'TRUE' }
VERSION : 1.0
   VAR_INPUT
      hardware_id : Port;   // hardware id
      operating_mode : USInt := 4;   // 0: RS232, 2: RS422, 4: RS485.
      baud : UDInt := 19200;   // Bits per sec.
   END_VAR
   VAR_OUTPUT
      Error : Bool;   // One or more errors in the whole application.
   END_VAR
   VAR_IN_OUT
      mb_query : "mb_query";
   END_VAR
   VAR
      conf : Struct   // Configuration that normal shouldn't need to be changed.
         parity : UInt := 2;   // 0=no-parity, 1=odd, 2=even.
         retries : USInt := 0;
         timeout : Time;   // Automatically calculated if set to zero. (T#0s)
      END_STRUCT;
      comm_load : Modbus_Comm_Load;
      master : Modbus_Master;
      buffer : "mb_internal_b";
      end : "mb_internal_e";
      comm_load_done : Bool;
      init_hw : Bool := true;
   END_VAR
   VAR CONSTANT
      INIT_QUERY : USInt := 2;
      EXEC_QUERY : USInt := 3;
      RECIVE_RESUALT : USInt := 4;
   END_VAR
BEGIN
   // Rexhip - Extended modbus library.
   // Please see top section of mb_query for more info.
   //
   // RTU master for S7-1500
   // 
   // This master blocks works for both S7-1200 and S7-1500. For S7-1200
   // it's recommended to use the other master block, mb_master_1200_ctrl
   // because it use less memory. Please read the documentation, before
   // dive into the code bellow.

   REGION Init
       IF #init_hw THEN
           // T#0s => Automatically adjust timeout.
           #comm_load.RESP_TO :=
           SEL(G := #conf.timeout = T#0s,
               IN0 := T_CONV(#conf.timeout),
               IN1 := UDINT_TO_UINT(4500000 / #baud));
       END_IF;
       // Initiate the hardware.
       #comm_load.RETRIES := #conf.retries;
       #comm_load.MODE := #operating_mode;
       #comm_load(REQ := #init_hw,
                  PORT := #hardware_id,
                  BAUD := #baud,
                  PARITY := #conf.parity, // Even is default.
                  RESP_TO := #comm_load.RESP_TO,
                  MB_DB := #master.MB_DB);
       #init_hw := false; // Hw init Finnised
       IF #comm_load.DONE THEN
           #comm_load_done := true;
       END_IF;

       IF #mb_query.z.run.state = #INIT_QUERY THEN
           // Modicon convention address conversion.
           "mb_internal_a"(mode104 := true,
                          Mode => #master.MODE,
                          Data_addr => #master.DATA_ADDR,
                          mb_query := #mb_query);

          // Copy buffer to a non optimiced memory area.
           IF #mb_query.z.run.write THEN
               #buffer.buffer := #mb_query.z.buffer;
           END_IF;

           IF #comm_load_done THEN
               #mb_query.z.run.state := #EXEC_QUERY;
           ELSE
               // Skip query exec. if init hw didn't go well.
               // The state RECIVE_RESUALT is inside mb_query.
               #mb_query.z.run.state := #RECIVE_RESUALT;
               #mb_query.stat.done := false;
               #mb_query.stat.error := true;
               #mb_query.stat.error_comm := true;
               #mb_query.stat.status := #comm_load.STATUS;
           END_IF;
       END_IF;
   END_REGION

   REGION Exec
       #master(REQ := #mb_query.z.run.state = #EXEC_QUERY
               AND NOT #master.BUSY,
               MB_ADDR := #mb_query.z.q.mb_addr,
               MODE := #master.MODE,
               DATA_ADDR := #master.DATA_ADDR,
               DATA_LEN := #mb_query.z.q.data_len,
               BUSY => #mb_query.stat.busy,
               DATA_PTR := #buffer.buffer);

       IF #mb_query.z.run.state = #EXEC_QUERY THEN
           #mb_query.stat.error := #master.ERROR;
           #mb_query.stat.done := #master.DONE;
           #mb_query.stat.status := #master.STATUS;
           "mb_internal_f"(buffer := #buffer, mb_query := #mb_query);
       END_IF;
   END_REGION

   // End is a comman FB for both tcp and rtu.
   #end(mb_query := #mb_query, Error => #Error);
END_FUNCTION_BLOCK

// folder: Library/Modbus/Core/Special

FUNCTION "mb_dataptr_eq_buffer" : Bool   // FC3, SCL
{ S7_Optimized_Access := 'TRUE' }